
Template "03_Three_Nav_Levels" 1280x800
   Gauge "gaugeDiagStateUpdate" at 566,2 size 50x50; CaptionText 'SIMATIC'
      on Change: "CheckDiagState"()
      ProcessValue <- "@DiagnosticsIndicatorTag"
   TextField "txtTitleBar" at 16,8 size 495x32; Text 'Application Name / Applikation'
   GraphicView "gfxNavigationIcon" at 1241,15 size 23x19; Picture "Hamburger_Icon"
   Button "btnNavigation" at 1224,0 size 56x48; TextOff 'Text'
      on Click: function_cf6f4242("GraphX_Slidein_Right", 1)
   TextField "txtStateHeadline" at 75,55 size 123x23; Text 'State / Status'
   TextField "txtRecipeHeadline" at 281,55 size 154x23; Text 'Current Recipe / Rezeptur'
   TextField "txtOperatorHeadline" at 527,55 size 129x23; Text 'Operator / Bediener'
   SymbolicIOField "ioState" at 75,72 size 119x30; TextOn '1'; TextOff '0'; TextList "Machine State"
      ProcessValue <- "CurrentMachineState"
   IOField "ioRecipe" at 281,72 size 158x30; FormatPattern ??????????????????????????????
      ProcessValue <- "CurrentRecipeName"
   IOField "ioOperator" at 527,72 size 126x30; FormatPattern ??????????????????
      ProcessValue <- "CurrentUserName"
   Button "btnState" at 202,56 size 40x40; TextOff '...'; PictureOff "More_Icon"
      on Click: "ShowOperatingModePopUp"()
   Button "btnRecipe" at 449,56 size 40x40; TextOff '...'; PictureOff "More_Icon"
      on Click: "ShowRecipePopUp"()
   Rectangle "rectState" at 0,48 size 56x56
      Appearance <- "CurrentMachineState"
   Rectangle "rectSystemDiagnosticsIndicator" at 1224,48 size 56x56
      Appearance <- "DiagState"
   GraphicIOField "gioDiagState" at 1236,60 size 32x32; PictureList "DiagState_3"
      ProcessValue <- "DiagState"
   Button "btnDiagState" at 1224,48 size 56x56; TextOff 'Text'
      on Click: ActivateScreen("30_Diagnostics", 0)
   Button "btnOperator" at 669,56 size 40x40; TextOff '...'; PictureOff "More_Icon"
      on Click: "ShowLoginPopUp"()
   TextField "txtOperatorHeadline_1" at 768,55 size 129x23; Text 'Date and Time / Bediener'
   Button "btnOperator_1" at 995,56 size 40x40; TextOff '...'; PictureOff "More_Icon"
   DateTimeField "Template_Date/time field_1" at 768,72 size 208x30
   Button "btnStartscreen" at 0,0 size 250x45; TextOff 'Text'
      on Click: "ActivateStartScreen"()
   Button "btnThirdLevel4btnOff1" at 0,104 size 56x163; TextOff 'Text'
   Button "btnThirdLevel4btnOff2" at 0,266 size 56x162; TextOff 'Text'
   Button "btnThirdLevel4btnOff3" at 0,427 size 56x163; TextOff 'Text'
   Button "btnThirdLevel4btnOff4" at 0,589 size 56x163; TextOff 'Text'
   Button "btnThirdLevel4btnOn1" at 0,266 size 56x161; TextOff 'Text'
      Visibility <- "ThirdLevelNavigationState"
   Button "btnThirdLevel4btnOn2" at 0,104 size 56x161; TextOff 'Text'
      Visibility <- "ThirdLevelNavigationState"
   Button "btnThirdLevel4btnOn3" at 0,428 size 56x161; TextOff 'Text'
      Visibility <- "ThirdLevelNavigationState"
   Button "btnThirdLevel4btnOn4" at 0,590 size 56x162; TextOff 'Text'
      Visibility <- "ThirdLevelNavigationState"
   Rectangle "rectIndicator4btnActive1" at 0,104 size 5x161
      Visibility <- "ThirdLevelNavigationState"
   Rectangle "rectIndicator4btnActive2" at 0,266 size 5x161
      Visibility <- "ThirdLevelNavigationState"
   Rectangle "rectIndicator4btnActive3" at 0,428 size 5x161
      Visibility <- "ThirdLevelNavigationState"
   Rectangle "rectIndicator4btnActive4" at 0,590 size 5x162
      Visibility <- "ThirdLevelNavigationState"
   Button "btnSubNavActive1" at 0,752 size 144x48; TextOff 'Overview / Übersicht'
      Visibility <- "SubNavigationState"
   Button "btnSubNavActive2" at 144,752 size 144x48; TextOff 'Module 1 / Modul 1'
      Visibility <- "SubNavigationState"
   Button "btnSubNavActive3" at 288,752 size 144x48; TextOff 'Module 2 / Modul 2'
      Visibility <- "SubNavigationState"
   Button "btnSubNavActive4" at 432,752 size 144x48; TextOff 'Module 3 / Modul 3'
      Visibility <- "SubNavigationState"
   Button "btnSubNavActive5" at 576,752 size 144x48; TextOff 'Module 4 / Modul 4'
      Visibility <- "SubNavigationState"
   Button "btnSubNavActive6" at 720,752 size 144x48; TextOff 'Module 5 / Modul 5'
      Visibility <- "SubNavigationState"
   Button "btnSubNavActive7" at 864,752 size 144x48; TextOff 'Module 6 / Modul 5'
      Visibility <- "SubNavigationState"
   Rectangle "rectIndicatorActive1" at 0,795 size 144x5
      Visibility <- "SubNavigationState"
   Rectangle "rectIndicatorActive2" at 144,795 size 144x5
      Visibility <- "SubNavigationState"
   Rectangle "rectIndicatorActive3" at 288,795 size 144x5
      Visibility <- "SubNavigationState"
   Rectangle "rectIndicatorActive4" at 432,795 size 144x5
      Visibility <- "SubNavigationState"
   Rectangle "rectIndicatorActive5" at 576,795 size 144x5
      Visibility <- "SubNavigationState"
   Rectangle "rectIndicatorActive6" at 720,795 size 144x5
      Visibility <- "SubNavigationState"
   Rectangle "rectIndicatorActive7" at 864,795 size 144x5
      Visibility <- "SubNavigationState"
   GraphicView "gfxPrevScreenIcon" at 1240,763 size 24x24; Picture "PrevScreen_Icon"
   Button "btnSubNav1" at 0,752 size 144x48; TextOff 'Overview / Übersicht'
      on Click: SetTag("SubNavigationState", 1)
   Button "btnSubNav2" at 144,752 size 144x48; TextOff 'Module 1 / Modul 1'
      on Click: SetTag("SubNavigationState", 2)
   Button "btnSubNav3" at 288,752 size 144x48; TextOff 'Module 2 / Modul 2'
      on Click: SetTag("SubNavigationState", 3)
   Button "btnSubNav4" at 432,752 size 144x48; TextOff 'Module 3 / Modul 3'
      on Click: SetTag("SubNavigationState", 4)
   Button "btnSubNav5" at 576,752 size 144x48; TextOff 'Module 4 / Modul 4'
      on Click: SetTag("SubNavigationState", 5)
   Button "btnSubNav6" at 720,752 size 144x48; TextOff 'Module 5 / Modul 5'
      on Click: SetTag("SubNavigationState", 6)
   Button "btnSubNav7" at 864,752 size 144x48; TextOff 'Module 6 / Modul 5'
      on Click: SetTag("SubNavigationState", 7)
   Button "btnPreviousScreen" at 1224,751 size 56x48; TextOff 'Text'
      on Click: function_efd93a16()

Template "03_Three_Nav_Levels_w_OptionPanel" 1280x800
   Gauge "gaugeDiagStateUpdate" at 566,2 size 50x50; CaptionText 'SIMATIC'
      on Change: "CheckDiagState"()
      ProcessValue <- "@DiagnosticsIndicatorTag"
   TextField "txtTitleBar" at 16,8 size 495x32; Text 'Application Name / Applikation'
   GraphicView "gfxNavigationIcon" at 1241,15 size 23x19; Picture "Hamburger_Icon"
   Button "btnNavigation" at 1224,0 size 56x48; TextOff 'Text'
      on Click: function_cf6f4242("GraphX_Slidein_Right", 1)
   TextField "txtStateHeadline" at 75,55 size 123x23; Text 'State / Status'
   TextField "txtRecipeHeadline" at 281,55 size 154x23; Text 'Current Recipe / Rezeptur'
   TextField "txtOperatorHeadline" at 527,55 size 129x23; Text 'Operator / Bediener'
   SymbolicIOField "ioState" at 75,72 size 119x30; TextOn '1'; TextOff '0'; TextList "Machine State"
      ProcessValue <- "CurrentMachineState"
   IOField "ioRecipe" at 281,72 size 158x30; FormatPattern ??????????????????????????????
      ProcessValue <- "CurrentRecipeName"
   IOField "ioOperator" at 527,72 size 126x30; FormatPattern ??????????????????
      ProcessValue <- "CurrentUserName"
   Button "btnState" at 202,56 size 40x40; TextOff '...'; PictureOff "More_Icon"
      on Click: "ShowOperatingModePopUp"()
   Button "btnRecipe" at 449,56 size 40x40; TextOff '...'; PictureOff "More_Icon"
      on Click: "ShowRecipePopUp"()
   Rectangle "rectState" at 0,48 size 56x56
      Appearance <- "CurrentMachineState"
   Rectangle "rectSystemDiagnosticsIndicator" at 1224,48 size 56x56
      Appearance <- "DiagState"
   GraphicIOField "gioDiagState" at 1236,60 size 32x32; PictureList "DiagState_3"
      ProcessValue <- "DiagState"
   Button "btnDiagState" at 1224,48 size 56x56; TextOff 'Text'
      on Click: ActivateScreen("30_Diagnostics", 0)
   Button "btnOperator" at 669,56 size 40x40; TextOff '...'; PictureOff "More_Icon"
      on Click: "ShowLoginPopUp"()
   TextField "txtOperatorHeadline_1" at 768,55 size 129x23; Text 'Date and Time / Bediener'
   Button "btnOperator_1" at 995,56 size 40x40; TextOff '...'; PictureOff "More_Icon"
   DateTimeField "Template_Date/time field_1" at 768,72 size 208x30
   Button "btnStartscreen" at 0,0 size 250x45; TextOff 'Text'
      on Click: "ActivateStartScreen"()
   Button "btnThirdLevel4btnOff1" at 0,104 size 56x163; TextOff 'Text'
   Button "btnThirdLevel4btnOff2" at 0,266 size 56x162; TextOff 'Text'
   Button "btnThirdLevel4btnOff3" at 0,427 size 56x163; TextOff 'Text'
   Button "btnThirdLevel4btnOff4" at 0,589 size 56x163; TextOff 'Text'
   Button "btnThirdLevel4btnOn1" at 0,266 size 56x161; TextOff 'Text'
      Visibility <- "ThirdLevelNavigationState"
   Button "btnThirdLevel4btnOn2" at 0,104 size 56x161; TextOff 'Text'
      Visibility <- "ThirdLevelNavigationState"
   Button "btnThirdLevel4btnOn3" at 0,428 size 56x161; TextOff 'Text'
      Visibility <- "ThirdLevelNavigationState"
   Button "btnThirdLevel4btnOn4" at 0,590 size 56x162; TextOff 'Text'
      Visibility <- "ThirdLevelNavigationState"
   Rectangle "rectIndicator4btnActive1" at 0,104 size 5x161
      Visibility <- "ThirdLevelNavigationState"
   Rectangle "rectIndicator4btnActive2" at 0,266 size 5x161
      Visibility <- "ThirdLevelNavigationState"
   Rectangle "rectIndicator4btnActive3" at 0,428 size 5x161
      Visibility <- "ThirdLevelNavigationState"
   Rectangle "rectIndicator4btnActive4" at 0,590 size 5x162
      Visibility <- "ThirdLevelNavigationState"
   Button "btnOptionbtn1" at 1224,104 size 56x648; TextOff 'Text'; PictureOn "ManFunctions_Off"; PictureOff "ManFunctions_Off"
      on Click: "ShowOptionPanelPopUp"()
   GraphicView "gfxPrevScreenIcon" at 1240,763 size 24x24; Picture "PrevScreen_Icon"
   Button "btnSubNav1" at 0,752 size 144x48; TextOff 'Overview / Übersicht'
      on Click: SetTag("SubNavigationState", 1)
   Button "btnSubNav2" at 144,752 size 144x48; TextOff 'Module 1 / Modul 1'
      on Click: SetTag("SubNavigationState", 2)
   Button "btnSubNav3" at 288,752 size 144x48; TextOff 'Module 2 / Modul 2'
      on Click: SetTag("SubNavigationState", 3)
   Button "btnSubNav4" at 432,752 size 144x48; TextOff 'Module 3 / Modul 3'
      on Click: SetTag("SubNavigationState", 4)
   Button "btnSubNav5" at 576,752 size 144x48; TextOff 'Module 4 / Modul 4'
      on Click: SetTag("SubNavigationState", 5)
   Button "btnSubNav6" at 720,752 size 144x48; TextOff 'Module 5 / Modul 5'
      on Click: SetTag("SubNavigationState", 6)
   Button "btnSubNav7" at 864,752 size 144x48; TextOff 'Module 6 / Modul 5'
      on Click: SetTag("SubNavigationState", 7)
   Button "btnPreviousScreen" at 1224,751 size 56x48; TextOff 'Text'
      on Click: function_efd93a16()
   Button "btnSubNavActive1" at 0,752 size 144x48; TextOff 'Overview / Übersicht'
      Visibility <- "SubNavigationState"
   Button "btnSubNavActive2" at 144,752 size 144x48; TextOff 'Module 1 / Modul 1'
      Visibility <- "SubNavigationState"
   Button "btnSubNavActive3" at 288,752 size 144x48; TextOff 'Module 2 / Modul 2'
      Visibility <- "SubNavigationState"
   Button "btnSubNavActive4" at 432,752 size 144x48; TextOff 'Module 3 / Modul 3'
      Visibility <- "SubNavigationState"
   Button "btnSubNavActive5" at 576,752 size 144x48; TextOff 'Module 4 / Modul 4'
      Visibility <- "SubNavigationState"
   Button "btnSubNavActive6" at 720,752 size 144x48; TextOff 'Module 5 / Modul 5'
      Visibility <- "SubNavigationState"
   Button "btnSubNavActive7" at 864,752 size 144x48; TextOff 'Module 6 / Modul 5'
      Visibility <- "SubNavigationState"
   Rectangle "rectIndicatorActive1" at 0,795 size 144x5
      Visibility <- "SubNavigationState"
   Rectangle "rectIndicatorActive2" at 144,795 size 144x5
      Visibility <- "SubNavigationState"
   Rectangle "rectIndicatorActive3" at 288,795 size 144x5
      Visibility <- "SubNavigationState"
   Rectangle "rectIndicatorActive4" at 432,795 size 144x5
      Visibility <- "SubNavigationState"
   Rectangle "rectIndicatorActive5" at 576,795 size 144x5
      Visibility <- "SubNavigationState"
   Rectangle "rectIndicatorActive6" at 720,795 size 144x5
      Visibility <- "SubNavigationState"
   Rectangle "rectIndicatorActive7" at 864,795 size 144x5
      Visibility <- "SubNavigationState"

Template "02_Settings" 1280x800
   Button "btnSubNav1" at 0,184 size 136x56; TextOn 'Display'; TextOff 'Display'
      on Click: SetTag("SubNavigationState", 1)
   GraphicView "gfxRuntimeStop" at 57,763 size 23x28; Picture "Power_dark"
   Button "btnRuntimeStop" at 0,751 size 136x48; TextOff 'Text'
      on Click: StopRuntime(0); SetBit("DB_UDP_COMM_PLC_TO_PC_TUSEND_DB_TUSEND_REQ")
   Button "btnSubNavActive1" at 0,184 size 136x56; TextOn 'Display'; TextOff 'Display'
      Visibility <- "SubNavigationState"
   Rectangle "rectIndicatorActive1" at 0,184 size 5x56
      Visibility <- "SubNavigationState"
   Gauge "gaugeDiagStateUpdate" at 566,2 size 50x50; CaptionText 'SIMATIC'
      on Change: "CheckDiagState"()
      ProcessValue <- "@DiagnosticsIndicatorTag"
   TextField "txtTitleBar" at 16,8 size 613x32; Text 'Application Name / Applikation'
   GraphicView "gfxNavigationIcon" at 1241,15 size 23x19; Picture "Hamburger_Icon"
   Button "btnNavigation" at 1224,0 size 56x48; TextOff 'Text'
      on Click: function_cf6f4242("GraphX_Slidein_Right", 1)
   Button "btnStartscreen" at 0,0 size 387x45; TextOff 'Text'
      on Click: "ActivateStartScreen"()
   TextField "txtStateHeadline" at 75,55 size 123x23; Text 'State / Status'
   TextField "txtRecipeHeadline" at 281,55 size 154x23; Text 'Current Recipe / Rezeptur'
   TextField "txtOperatorHeadline" at 527,55 size 129x23; Text 'Operator / Bediener'
   SymbolicIOField "ioState" at 75,72 size 119x30; TextOn '1'; TextOff '0'; TextList "Machine State"
      ProcessValue <- "CurrentMachineState"
   IOField "ioRecipe" at 281,72 size 158x30; FormatPattern ??????????????????????????????
      ProcessValue <- "CurrentRecipeName"
   IOField "ioOperator" at 527,72 size 126x30; FormatPattern ??????????????????
      ProcessValue <- "CurrentUserName"
   Button "btnState" at 202,56 size 40x40; TextOff '...'; PictureOff "More_Icon"
      on Click: "ShowOperatingModePopUp"()
   Button "btnRecipe" at 449,56 size 40x40; TextOff '...'; PictureOff "More_Icon"
      on Click: "ShowRecipePopUp"()
   Rectangle "rectState" at 0,48 size 56x56
      Appearance <- "CurrentMachineState"
   Rectangle "rectSystemDiagnosticsIndicator" at 1224,48 size 56x56
      Appearance <- "DiagState"
   GraphicIOField "gioDiagState" at 1236,60 size 32x32; PictureList "DiagState_3"
      ProcessValue <- "DiagState"
   Button "btnDiagState" at 1224,48 size 56x56; TextOff 'Text'
      on Click: ActivateScreen("30_Diagnostics", 0)
   Button "btnOperator" at 669,56 size 40x40; TextOff '...'; PictureOff "More_Icon"
      on Click: "ShowLoginPopUp"()
   TextField "txtOperatorHeadline_1" at 768,55 size 129x23; Text 'Date and Time / Bediener'
   Button "btnOperator_1" at 995,56 size 40x40; TextOff '...'; PictureOff "More_Icon"
   DateTimeField "Template_Date/time field_1" at 768,72 size 208x30

PopupScreen "Template_Logon" 320x352
   on ClearScreen: ResetBit("PopUpBackground")
   on GenerateScreen: SetBit("PopUpBackground")
   TextField "Template_Text field_1" at 16,0 size 215x40; Text 'Login'
   Button "Button_2" at 16,240 size 288x40; TextOn 'LOGIN / ANMELDEN'; TextOff 'LOGIN / ANMELDEN'
      on Click: function_a9b89908("Password", "UserName"); function_efd93a16("Template_Logon", 0, 0, 0, -1, 1)
   IOField "I/O field_1" at 16,84 size 288x40; FormatPattern ??????????????????????????????
      ProcessValue <- "UserName"
   TextField "Text field_1" at 16,56 size 288x24; Text 'User Name / Name'
   IOField "I/O field_2" at 16,168 size 288x40; FormatPattern ??????????????????????????????
      ProcessValue <- "Password"
   TextField "Text field_2" at 16,140 size 288x24; Text 'Password / Passwort'
   Button "Button_1" at 16,296 size 288x40; TextOn 'CLOSE / SCHLIESSEN'; TextOff 'CLOSE / SCHLIESSEN'
      on Click: function_efd93a16("Template_Logon", 0, 0, 0, -1, 1)
      on Press: function_b14e0dd5("ButtonDown", 0)
      Appearance <- "ButtonDown"

PopupScreen "Template_Logon_Logoff" 320x352
   on ClearScreen: ResetBit("PopUpBackground")
   on GenerateScreen: SetBit("PopUpBackground")
   TextField "Template_Text field_1" at 16,0 size 215x40; Text 'Login'
   Button "Button_2" at 16,240 size 136x40; TextOn 'LOG OFF / ABMELDEN'; TextOff 'LOG OFF / ABMELDEN'
      on Click: function_f23ef4c9()
   IOField "I/O field_1" at 16,84 size 288x40; FormatPattern ??????????????????????????????
      ProcessValue <- "UserName"
   TextField "Text field_1" at 16,56 size 288x24; Text 'User Name / Name'
   IOField "I/O field_2" at 16,168 size 288x40; FormatPattern ??????????????????????????????
      ProcessValue <- "Password"
   TextField "Text field_2" at 16,140 size 288x24; Text 'Password / Passwort'
   Button "Button_1" at 16,296 size 288x40; TextOn 'CLOSE / SCHLIESSEN'; TextOff 'CLOSE / SCHLIESSEN'
      on Click: function_efd93a16("Template_Logon_Logoff", 0, 0, 0, -1, 1)
      on Press: function_b14e0dd5("ButtonDown", 0)
      Appearance <- "ButtonDown"
   Button "Button_3" at 168,240 size 136x40; TextOn 'LOGIN / ANMELDEN'; TextOff 'LOGIN / ANMELDEN'
      on Click: function_a9b89908("Password", "UserName"); function_efd93a16("Template_Logon_Logoff", 0, 0, 0, -1, 1)

PopupScreen "Template_Operating_Mode" 424x360
   on ClearScreen: ResetBit("PopUpBackground")
   on GenerateScreen: SetBit("PopUpBackground")
   TextField "Template_Text field_1" at 14,0 size 336x40; Text 'Operating Mode / Betriebsmodus'
   Button "Button_1" at 80,304 size 260x40; TextOn 'CLOSE / SCHLIESSEN'; TextOff 'CLOSE / SCHLIESSEN'
      on Click: function_efd93a16("Template_Operating_Mode", 0, 0, 0, -1, 1)
      on Press: function_b14e0dd5("ButtonDown", 0)
      Appearance <- "ButtonDown"
   Button "Button_2" at 352,66 size 40x40; TextOff 'Text'; PictureOff "More_Icon"; PictureOn "More_Icon"
   Button "Button_3" at 352,130 size 40x40; TextOff 'Text'; PictureOn "More_Icon"; PictureOff "More_Icon"
   Button "Button_4" at 28,210 size 82x48; TextOff 'Start'
   Button "Button_5" at 123,210 size 82x48; TextOff 'Stop'
   Button "Button_6" at 218,210 size 82x48; TextOff 'Reset'
   Button "Button_7" at 314,210 size 82x48; TextOff 'Hold'
   TextField "txtParameter7_3" at 32,63 size 163x24; Text 'Current Mode'
   IOField "ioParameter17_3" at 32,81 size 301x40; FormatPattern ?????????????????????????
   TextField "txtParameter7_1" at 32,127 size 163x24; Text 'Current State'
   IOField "ioParameter17_1" at 32,145 size 301x40; FormatPattern ?????????????????????????

PopupScreen "Template_Recipe" 700x420
   on ClearScreen: ResetBit("PopUpBackground")
   on GenerateScreen: SetBit("PopUpBackground")
   TextField "Template_Text field_1" at 14,0 size 500x40; Text 'Recipe / Rezeptur'
   Button "Button_1" at 220,364 size 260x40; TextOn 'CLOSE / SCHLIESSEN'; TextOff 'CLOSE / SCHLIESSEN'
      on Click: function_efd93a16("Template_Recipe", 0, 0, 0, -1, 1)
      on Press: function_b14e0dd5("ButtonDown", 0)
      Appearance <- "ButtonDown"

PopupScreen "OptionPanel_4_Buttons" 390x648
   Button "btnCloseOptionPanel" at 0,0 size 40x648; TextOff 'CLOSE'; PictureOff "Jog_Forward"
      on Press: function_efd93a16("OptionPanel_4_Buttons", 0, 0, 0, 2, 2)
   TextField "txtOptionPanel" at 108,16 size 260x40; Text 'Option Panel Title / Titel Option Panel'
   Button "btnOption1" at 80,72 size 240x40; TextOff 'Option 1 / Move to Home Position'
   Button "btnOption2" at 80,128 size 240x40; TextOff 'Option 2 / Move to Home Position'
   Button "btnOption3" at 80,184 size 240x40; TextOff 'Option 3 / RESET'
   Button "btnOption4" at 80,240 size 240x40; TextOff 'Option 4 / RESET'
   GraphicView "gvOptionPanel" at 80,30 size 18x12; Picture "ManFunctions_Off"

SlideinScreen "GraphX_Slidein_Left" 220x800
   Button "Button_1" at 15,220 size 188x72; TextOff 'RESET'
      on Press: SetBit("DB_HMI_Varjenje_ResetWithWC")
      on Release: ResetBit("DB_HMI_Varjenje_ResetWithWC")
   Button "Button_2" at 15,308 size 188x72; TextOff 'RESET + ZVAR'
   SymbolicIOField "Symbolic I/O field_1" at 10,437 size 201x29; TextOff '0'; TextOn '1'; TextList "BOSH"
      ProcessValue <- "StatusCode"
   TextField "Text field_1" at 22,267 size 176x23; Text 'Reset varilnika z WC'
   TextField "Text field_2" at 23,355 size 176x23; Text 'Reset varilnika z zvarom'
   TextField "Text field_3" at 10,414 size 176x23; Text 'STATUS VARILNIKA:'

SlideinScreen "GraphX_Slidein_Right" 220x800
   Button "Button_1" at 0,78 size 220x60; TextOn 'Menu Item 1'; TextOff 'Startscreen / Menu Item 1'
      on Click: SetTag("MainNavigationState", 1); ActivateScreen("10_Startup", 0)
      Appearance <- "MainNavigationState"
   Button "Button_2" at 0,140 size 220x60; TextOn 'Menu Item 2'; TextOff 'Lista napak / Menu Item 2'
      on Click: SetTag("MainNavigationState", 2); ActivateScreen("20_Messages", 0)
      Appearance <- "MainNavigationState"
   Button "Button_3" at 0,201 size 220x60; TextOn 'Menu Item 3'; TextOff 'Diagnostika / Menu Item 3'
      on Click: SetTag("MainNavigationState", 3); ActivateScreen("30_Diagnostics", 0)
      Appearance <- "MainNavigationState"
   Rectangle "Rectangle_1" at 214,78 size 6x60
      Visibility <- "MainNavigationState"
   Rectangle "Rectangle_2" at 214,140 size 6x60
      Visibility <- "MainNavigationState"
   Rectangle "Rectangle_3" at 214,201 size 6x60
      Visibility <- "MainNavigationState"
   Button "Button_4" at 0,262 size 220x60; TextOn 'Menu Item 4'; TextOff 'HMI / Menu Item 4'
      on Click: SetTag("MainNavigationState", 4); ActivateScreen("40_Settings", 0)
      Appearance <- "MainNavigationState"
   Rectangle "Rectangle_4" at 214,262 size 6x60
      Visibility <- "MainNavigationState"
   Button "Button_5" at 0,323 size 220x60; TextOn 'Menu Item 4'; TextOff 'Nastavitve / Menu Item 4'; Authorization "User administration"
      on Click: SetTag("MainNavigationState", 5); ActivateScreen("106_Rocno_postaja6", 0); SetTag("ThirdLevelNavigationState", 6)
      Appearance <- "MainNavigationState"
   Rectangle "Rectangle_5" at 214,323 size 6x60
      Visibility <- "MainNavigationState"
   Button "Button_6" at 0,740 size 220x60; TextOn 'Menu Item 4'; TextOff 'Izklop stroja / Menu Item 4'
      on Click: SetTag("MainNavigationState", 10)
      Appearance <- "MainNavigationState"
   Rectangle "Rectangle_6" at 212,738 size 6x60
      Visibility <- "MainNavigationState"
   GraphicView "Graphic view_1" at 155,750 size 47x37; Picture "ExitRuntime_TP1200_Comfort_TR"
   Button "btnRuntimeStop" at 0,732 size 219x68; TextOff 'Text'
      on Click: StopRuntime(0); SetBit("DB_UDP_COMM_PLC_TO_PC_TUSEND_DB_TUSEND_REQ")

screen "10_Startup" 1280x800, template "01_One_Nav_Level"
   on GenerateScreen: "GetStartScreenName"(); "CheckCurrentUserName"()
   GraphicView "Graphic view_2" at 0,0 size 1280x800; Picture "PopUpBackground"
      Visibility <- "PopUpBackground"
   TextField "Text field_1" at 944,179 size 67x25; Text 'SERVO'
   Rectangle "Rectangle_1" at 1082,179 size 23x23
      Appearance <- "FB_AKD_DB_elektroda_o_BerrStatus"
   Rectangle "Rectangle_3" at 1152,179 size 23x23
      Appearance <- "FB_AKD_DB_RezanjePodajanje_o_BerrStatus"
   TextField "Text field_7" at 944,233 size 99x25; Text 'VARJENJE'
   TextField "Text field_2" at 1186,263 size 19x25; Text 'Q'
   TextField "Text field_3" at 1189,292 size 16x25; Text 'T'
   Rectangle "Rectangle_5" at 1213,263 size 23x23
      Appearance <- "FB_IOL_IFM_SV_DB_oPretokOK"
   Rectangle "Rectangle_6" at 1213,292 size 23x23
      Appearance <- "FB_IOL_IFM_SV_DB_oTempOK"
   TextField "Text field_4" at 1175,235 size 58x25; Text 'VODA'
   TextField "Text field_9" at 944,354 size 197x25; Text 'PRISOTNOST TRAKU'
   IOField "I/O field_1" at 937,742 size 129x32; FormatPattern 99999; Unit  l/min
      ProcessValue <- "FB_IOL_IFM_SV_DB_uPretok"
   IOField "I/O field_2" at 1074,742 size 84x32; FormatPattern 99.9; Unit  °C
      ProcessValue <- "FB_IOL_IFM_SV_DB_fTemperatura"
   IOField "I/O field_3" at 1167,742 size 98x32; FormatPattern 99.9; Unit  bar
      ProcessValue <- "FB_Lin_FESTO_PNEVMATIKA_PRITISK_Q_izhod"
   Rectangle "Rectangle_8" at 1213,354 size 23x23
      Appearance <- "StatusPrisotnostiTraku"
   Rectangle "Rectangle_10" at 1117,179 size 23x23
      Appearance <- "FB_AKD_VrtenjeKroznika_o_BerrStatus"
   GraphicView "Graphic view_1" at 91,111 size 735x664; Picture "S1054-900-001"
   Rectangle "Rectangle_15" at 87,379 size 176x15
      Appearance <- "DB_PODATKI_KROZNA_MIZA_IzdelekPrisotenArray{7}"
   Polygon "Polygon_1" at 248,285 size 51x51
      Appearance <- "DB_PODATKI_KROZNA_MIZA_IzdelekPrisoten"
   Polygon "Polygon_2" at 160,197 size 139x139
      Appearance <- "DB_PODATKI_KROZNA_MIZA_IzdelekPrisotenArray{6}"
   Polygon "Polygon_3" at 344,120 size 15x78
      Appearance <- "DB_PODATKI_KROZNA_MIZA_StatusIzdelka{5}"
   Polygon "Polygon_4" at 342,194 size 16x116
      Appearance <- "DB_PODATKI_KROZNA_MIZA_IzdelekPrisotenArray{5}"
   Polygon "Polygon_5" at 482,195 size 59x61
      Appearance <- "DB_PODATKI_KROZNA_MIZA_StatusIzdelka{4}"
   Rectangle "Rectangle_16" at 544,377 size 68x18
      Appearance <- "DB_PODATKI_KROZNA_MIZA_StatusIzdelka{3}"
   Polygon "Polygon_6" at 481,518 size 60x59
      Appearance <- "DB_PODATKI_KROZNA_MIZA_StatusIzdelka{2}"
   Polygon "Polygon_7" at 403,245 size 90x89
      Appearance <- "DB_PODATKI_KROZNA_MIZA_IzdelekPrisotenArray{4}"
   Polygon "Polygon_8" at 429,377 size 60x19
      Appearance <- "DB_PODATKI_KROZNA_MIZA_IzdelekPrisotenArray{3}"
   Polygon "Polygon_9" at 403,439 size 54x51
      Appearance <- "DB_PODATKI_KROZNA_MIZA_IzdelekPrisotenArray{2}"
   Polygon "Polygon_10" at 344,464 size 15x66
      Appearance <- "DB_PODATKI_KROZNA_MIZA_IzdelekPrisotenArray{1}"
   Polygon "Polygon_11" at 342,579 size 17x68
      Appearance <- "DB_PODATKI_KROZNA_MIZA_StatusIzdelkaVarjenje{1}"